(* Logix 5000 project; controller NWGG 1756-L72 rev 35.12; software revision 35.00; part 15 of 19 *)
(* tags used below, declared in another part *)
   Air_Gates_Opened : BOOL;
   ALM_Air_Gate_Failed_Open_Bin17 : ALARM_DIGITAL;
   ALM_Air_Gate_Failed_Open_Bin18 : ALARM_DIGITAL;
   ALM_Air_Gate_Failed_Open_Bin19 : ALARM_DIGITAL;
   ALM_Air_Gate_Failed_Open_Bin20 : ALARM_DIGITAL;
   ALM_Air_Gate_Failed_Open_Bin21 : ALARM_DIGITAL;
   ALM_Air_Gate_Failed_Open_Bin22 : ALARM_DIGITAL;
   ALM_Air_Gate_Failed_Open_Bin23 : ALARM_DIGITAL;
   ALM_Air_Gate_Failed_Open_Bin24 : ALARM_DIGITAL;
   ALM_Air_Gate_Failed_Open_Bin25 : ALARM_DIGITAL;
   ALM_Air_Gate_Failed_Open_Bin26 : ALARM_DIGITAL;
   ALM_Air_Gate_Failed_Open_Bin27 : ALARM_DIGITAL;
   ALM_Air_Gate_Failed_Open_Bin28 : ALARM_DIGITAL;
   Auto_Stop_Clean : BOOL;
   Belt : udt_Motor[16];
   Belts_Ready : BOOL;
   Belts_Running : BOOL;
   Bin_Clean_Pause : BOOL;
   Bin_Loadout_Control : Loadout_Bin_Control[29];
   Bin_Transfer_Pause : BOOL;
   Bin_Treat_Pause : BOOL;
   Bins_Rqd : BOOL;
   ckIDX : DINT;
   Clean_Batch_Status : DINT;
   Clean_Bin_Gates_Opened : BOOL;
   Clean_Interlock : BOOL;
   Clean_Scale_Unavailable : BOOL;
   cntCleanTime : COUNTER;
   Concrete_Clean_Belts_Ready : BOOL;
   Concrete_Leg : udt_Motor;
   Current_Dist_List_IDX : DINT;
   Current_Transfer_Bin_From : BOOL[32];
   Current_Transfer_Bin_To : BOOL[32];
   IDX : DINT;
   Loadout_Bin : udt_Loadout_Bin[29];
   Loadout_K_Valve : udt_Loadout_K_Valve[2];
   Loop_Idx : DINT;
   Manual_Mode : BOOL;
   NA : BOOL;
   Pause_Load_By_Time : BOOL[32];
   Pause_Load_By_Weight : BOOL[32];
   Pause_Load_Expired : DINT[2];
   Pause_Load_Pre : DINT[2];
   Reversing_Belt_Bypass_Valve : BOOL;
   Reversing_Belt_Reversed : BOOL;
   Start_Clean_Belts_Enabled : BOOL;
   Steel_Rqd_Belts_Running : BOOL;
   Target_Weight : DINT[2];
   TMR_Max_Clean_Delay : TIMER;
   TMR_Max_Treat_Delay : TIMER;
   tmr_Pause_Load_Timer : TIMER[2];
   tmrCleanTime : TIMER;
   Transfer_Batch_Status : DINT;
   Transfer_From_IDX : DINT;
   Transfer_To_IDX : DINT;
   Treat_Batch_Status : DINT;
   Treat_Bin_Gates_Opened : BOOL;
   Treat_Bins_Open : BOOL;
   Treat_Scale_Unavailable : BOOL;
   Use_Concrete_Side_Clean : BOOL;
   Use_Steel_Side_Clean : BOOL;
   Use_Steel_Transfer_Bins : BOOL;
   I1_000_Bit02 : ALIAS FOR I1.2;
   I1_000_Bit03 : ALIAS FOR I1.3;
   I1_000_Bit04 : ALIAS FOR I1.4;
   I1_000_Bit06 : ALIAS FOR I1.6;
   I1_000_Bit07 : ALIAS FOR I1.7;
   I1_000_Bit09 : ALIAS FOR I1.9;
   I1_000_Bit10 : ALIAS FOR I1.10;
   I1_000_Bit12 : ALIAS FOR I1.12;
   I1_000_Bit13 : ALIAS FOR I1.13;
   I1_000_Bit15 : ALIAS FOR I1.15;
   I2_000_Bit00 : ALIAS FOR I2.0;
   I2_000_Bit03 : ALIAS FOR I2.3;
   I2_000_Bit06 : ALIAS FOR I2.6;
   I2_000_Bit09 : ALIAS FOR I2.9;
   I2_000_Bit12 : ALIAS FOR I2.12;
   I3_000_Bit00 : ALIAS FOR I3.0;
   I3_000_Bit03 : ALIAS FOR I3.3;
   I3_000_Bit06 : ALIAS FOR I3.6;
   I4_000_Bit09 : ALIAS FOR I4.9;
   I4_000_Bit10 : ALIAS FOR I4.10;
   I4_000_Bit12 : ALIAS FOR I4.12;
   I4_000_Bit13 : ALIAS FOR I4.13;
   I4_000_Bit14 : ALIAS FOR I4.14;
   I4_000_Bit15 : ALIAS FOR I4.15;
   O10_000_Bit00 : ALIAS FOR O10.0;
   O10_000_Bit01 : ALIAS FOR O10.1;
   O10_000_Bit02 : ALIAS FOR O10.2;
   O10_000_Bit03 : ALIAS FOR O10.3;
   O10_000_Bit04 : ALIAS FOR O10.4;
   O10_000_Bit05 : ALIAS FOR O10.5;
   O10_000_Bit06 : ALIAS FOR O10.6;
   O10_000_Bit07 : ALIAS FOR O10.7;
   O10_000_Bit08 : ALIAS FOR O10.8;
   O10_000_Bit09 : ALIAS FOR O10.9;
   O10_000_Bit10 : ALIAS FOR O10.10;
   O10_000_Bit11 : ALIAS FOR O10.11;
   O10_000_Bit12 : ALIAS FOR O10.12;
   O10_000_Bit13 : ALIAS FOR O10.13;
   O10_000_Bit14 : ALIAS FOR O10.14;
   O11_000_Bit00 : ALIAS FOR O11.0;
   O11_000_Bit01 : ALIAS FOR O11.1;
   O11_000_Bit02 : ALIAS FOR O11.2;
   O11_000_Bit03 : ALIAS FOR O11.3;
   O11_000_Bit04 : ALIAS FOR O11.4;
   O11_000_Bit05 : ALIAS FOR O11.5;
   O11_000_Bit06 : ALIAS FOR O11.6;
   O11_000_Bit07 : ALIAS FOR O11.7;
   O11_000_Bit08 : ALIAS FOR O11.8;
   O9_000_Bit03 : ALIAS FOR O9.3;
   O9_000_Bit04 : ALIAS FOR O9.4;
   O9_000_Bit05 : ALIAS FOR O9.5;
   O9_000_Bit06 : ALIAS FOR O9.6;
   O9_000_Bit07 : ALIAS FOR O9.7;
   O9_000_Bit08 : ALIAS FOR O9.8;
   O9_000_Bit09 : ALIAS FOR O9.9;
   O9_000_Bit10 : ALIAS FOR O9.10;
   O9_000_Bit11 : ALIAS FOR O9.11;
   O9_000_Bit12 : ALIAS FOR O9.12;
   O9_000_Bit13 : ALIAS FOR O9.13;
   O9_000_Bit14 : ALIAS FOR O9.14;
   Truck_Scales : udt_Truck_Scale[2];
(* SeedLoadoutMain, continued *)

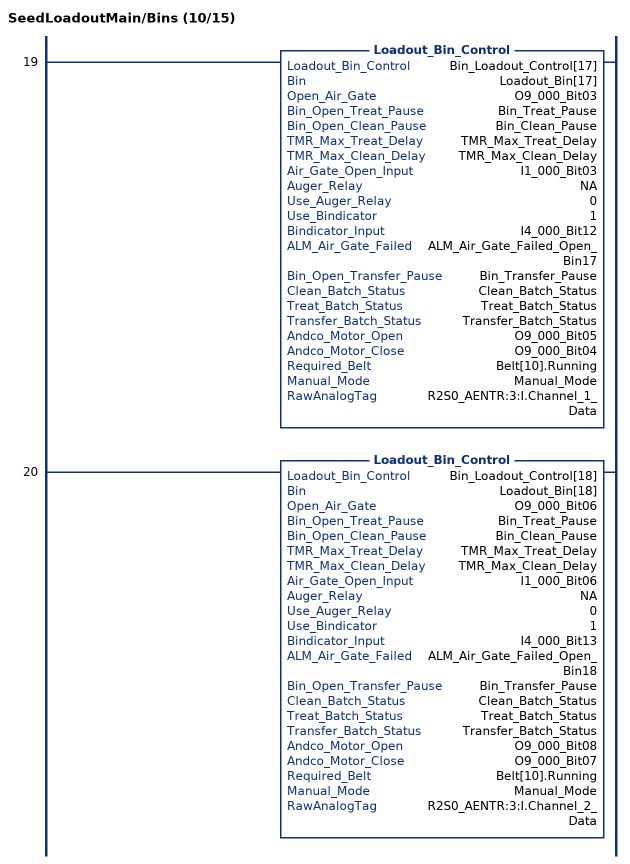
   19: Loadout_Bin_Control(Bin_Loadout_Control[17],Loadout_Bin[17],O9_000_Bit03,Bin_Treat_Pause,Bin_Clean_Pause,TMR_Max_Treat_Delay,TMR_Max_Clean_Delay,I1_000_Bit03,NA,0,1,I4_000_Bit12,ALM_Air_Gate_Failed_Open_Bin17,Bin_Transfer_Pause,Clean_Batch_Status,Treat_Batch_Status,Transfer_Batch_Status,O9_000_Bit05,O9_000_Bit04,Belt[10].Running,Manual_Mode,R2S0_AENTR:3:I.Channel_1_Data);
   20: Loadout_Bin_Control(Bin_Loadout_Control[18],Loadout_Bin[18],O9_000_Bit06,Bin_Treat_Pause,Bin_Clean_Pause,TMR_Max_Treat_Delay,TMR_Max_Clean_Delay,I1_000_Bit06,NA,0,1,I4_000_Bit13,ALM_Air_Gate_Failed_Open_Bin18,Bin_Transfer_Pause,Clean_Batch_Status,Treat_Batch_Status,Transfer_Batch_Status,O9_000_Bit08,O9_000_Bit07,Belt[10].Running,Manual_Mode,R2S0_AENTR:3:I.Channel_2_Data);
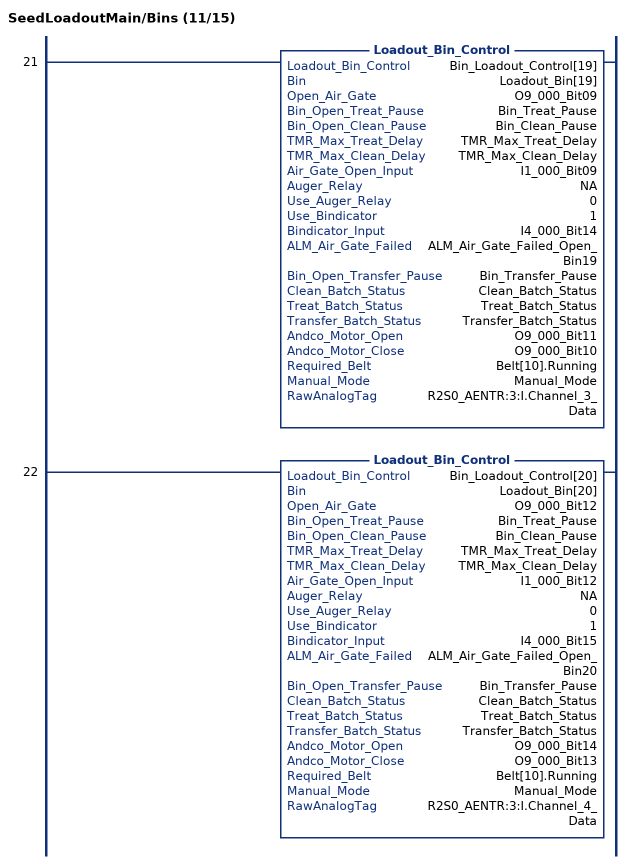
   21: Loadout_Bin_Control(Bin_Loadout_Control[19],Loadout_Bin[19],O9_000_Bit09,Bin_Treat_Pause,Bin_Clean_Pause,TMR_Max_Treat_Delay,TMR_Max_Clean_Delay,I1_000_Bit09,NA,0,1,I4_000_Bit14,ALM_Air_Gate_Failed_Open_Bin19,Bin_Transfer_Pause,Clean_Batch_Status,Treat_Batch_Status,Transfer_Batch_Status,O9_000_Bit11,O9_000_Bit10,Belt[10].Running,Manual_Mode,R2S0_AENTR:3:I.Channel_3_Data);
   22: Loadout_Bin_Control(Bin_Loadout_Control[20],Loadout_Bin[20],O9_000_Bit12,Bin_Treat_Pause,Bin_Clean_Pause,TMR_Max_Treat_Delay,TMR_Max_Clean_Delay,I1_000_Bit12,NA,0,1,I4_000_Bit15,ALM_Air_Gate_Failed_Open_Bin20,Bin_Transfer_Pause,Clean_Batch_Status,Treat_Batch_Status,Transfer_Batch_Status,O9_000_Bit14,O9_000_Bit13,Belt[10].Running,Manual_Mode,R2S0_AENTR:3:I.Channel_4_Data);
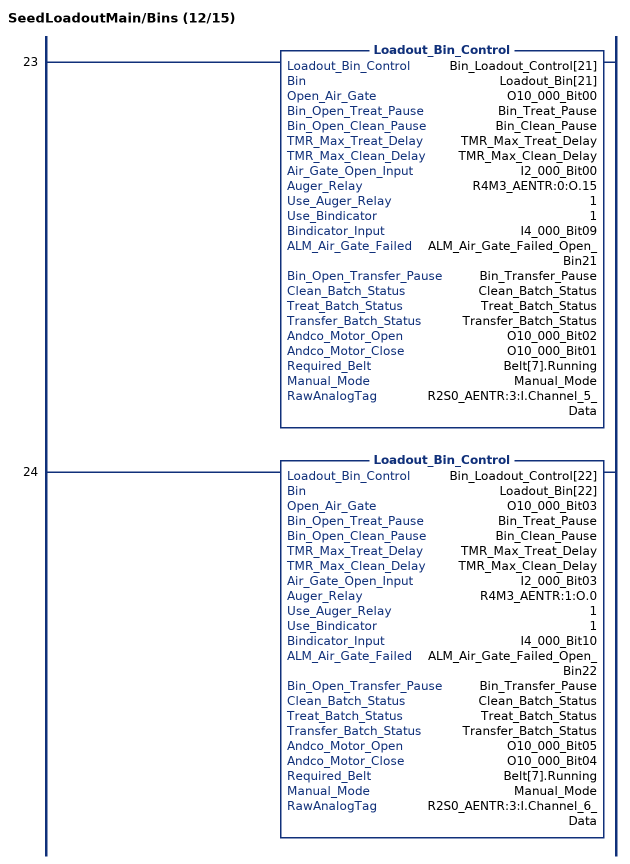
   23: Loadout_Bin_Control(Bin_Loadout_Control[21],Loadout_Bin[21],O10_000_Bit00,Bin_Treat_Pause,Bin_Clean_Pause,TMR_Max_Treat_Delay,TMR_Max_Clean_Delay,I2_000_Bit00,R4M3_AENTR:0:O.15,1,1,I4_000_Bit09,ALM_Air_Gate_Failed_Open_Bin21,Bin_Transfer_Pause,Clean_Batch_Status,Treat_Batch_Status,Transfer_Batch_Status,O10_000_Bit02,O10_000_Bit01,Belt[7].Running,Manual_Mode,R2S0_AENTR:3:I.Channel_5_Data);
   24: Loadout_Bin_Control(Bin_Loadout_Control[22],Loadout_Bin[22],O10_000_Bit03,Bin_Treat_Pause,Bin_Clean_Pause,TMR_Max_Treat_Delay,TMR_Max_Clean_Delay,I2_000_Bit03,R4M3_AENTR:1:O.0,1,1,I4_000_Bit10,ALM_Air_Gate_Failed_Open_Bin22,Bin_Transfer_Pause,Clean_Batch_Status,Treat_Batch_Status,Transfer_Batch_Status,O10_000_Bit05,O10_000_Bit04,Belt[7].Running,Manual_Mode,R2S0_AENTR:3:I.Channel_6_Data);
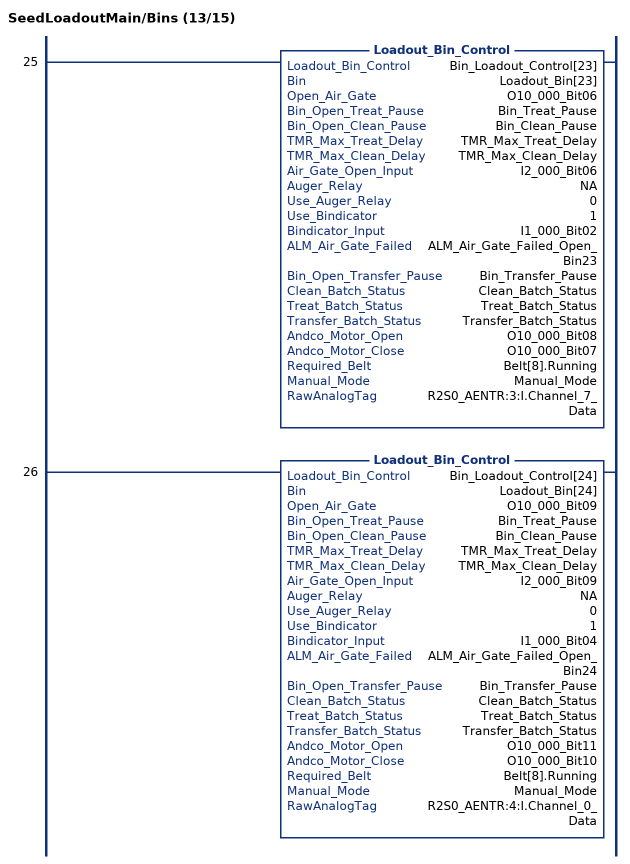
   25: Loadout_Bin_Control(Bin_Loadout_Control[23],Loadout_Bin[23],O10_000_Bit06,Bin_Treat_Pause,Bin_Clean_Pause,TMR_Max_Treat_Delay,TMR_Max_Clean_Delay,I2_000_Bit06,NA,0,1,I1_000_Bit02,ALM_Air_Gate_Failed_Open_Bin23,Bin_Transfer_Pause,Clean_Batch_Status,Treat_Batch_Status,Transfer_Batch_Status,O10_000_Bit08,O10_000_Bit07,Belt[8].Running,Manual_Mode,R2S0_AENTR:3:I.Channel_7_Data);
   26: Loadout_Bin_Control(Bin_Loadout_Control[24],Loadout_Bin[24],O10_000_Bit09,Bin_Treat_Pause,Bin_Clean_Pause,TMR_Max_Treat_Delay,TMR_Max_Clean_Delay,I2_000_Bit09,NA,0,1,I1_000_Bit04,ALM_Air_Gate_Failed_Open_Bin24,Bin_Transfer_Pause,Clean_Batch_Status,Treat_Batch_Status,Transfer_Batch_Status,O10_000_Bit11,O10_000_Bit10,Belt[8].Running,Manual_Mode,R2S0_AENTR:4:I.Channel_0_Data);
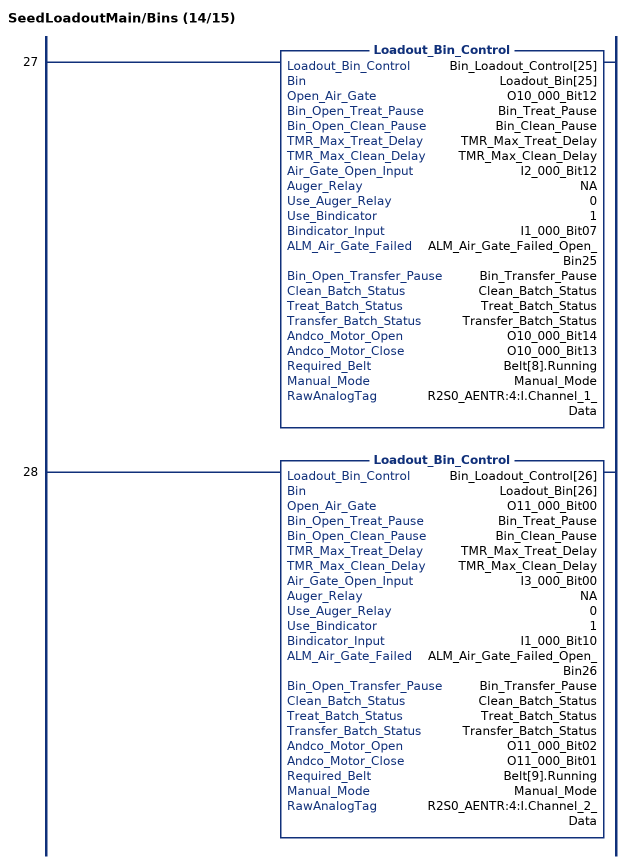
   27: Loadout_Bin_Control(Bin_Loadout_Control[25],Loadout_Bin[25],O10_000_Bit12,Bin_Treat_Pause,Bin_Clean_Pause,TMR_Max_Treat_Delay,TMR_Max_Clean_Delay,I2_000_Bit12,NA,0,1,I1_000_Bit07,ALM_Air_Gate_Failed_Open_Bin25,Bin_Transfer_Pause,Clean_Batch_Status,Treat_Batch_Status,Transfer_Batch_Status,O10_000_Bit14,O10_000_Bit13,Belt[8].Running,Manual_Mode,R2S0_AENTR:4:I.Channel_1_Data);
   28: Loadout_Bin_Control(Bin_Loadout_Control[26],Loadout_Bin[26],O11_000_Bit00,Bin_Treat_Pause,Bin_Clean_Pause,TMR_Max_Treat_Delay,TMR_Max_Clean_Delay,I3_000_Bit00,NA,0,1,I1_000_Bit10,ALM_Air_Gate_Failed_Open_Bin26,Bin_Transfer_Pause,Clean_Batch_Status,Treat_Batch_Status,Transfer_Batch_Status,O11_000_Bit02,O11_000_Bit01,Belt[9].Running,Manual_Mode,R2S0_AENTR:4:I.Channel_2_Data);
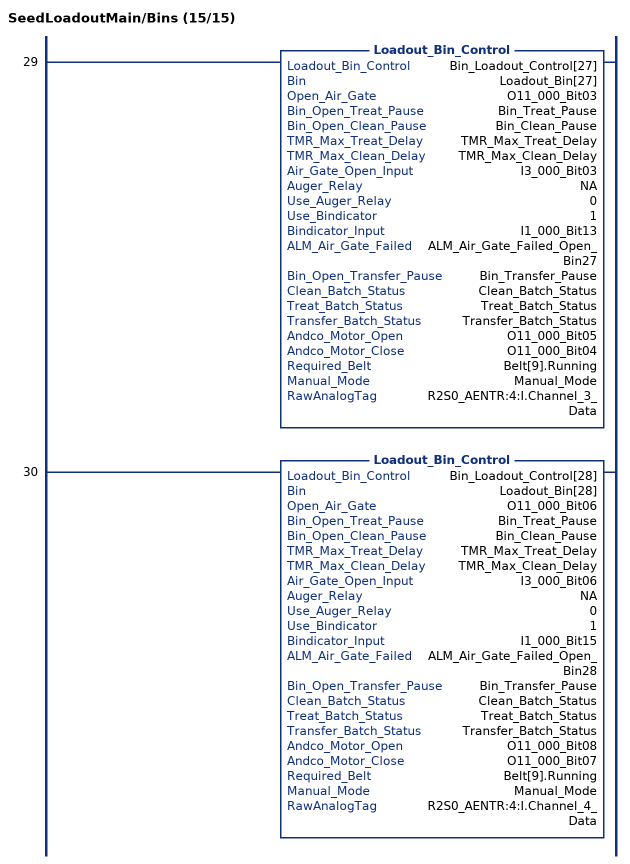
   29: Loadout_Bin_Control(Bin_Loadout_Control[27],Loadout_Bin[27],O11_000_Bit03,Bin_Treat_Pause,Bin_Clean_Pause,TMR_Max_Treat_Delay,TMR_Max_Clean_Delay,I3_000_Bit03,NA,0,1,I1_000_Bit13,ALM_Air_Gate_Failed_Open_Bin27,Bin_Transfer_Pause,Clean_Batch_Status,Treat_Batch_Status,Transfer_Batch_Status,O11_000_Bit05,O11_000_Bit04,Belt[9].Running,Manual_Mode,R2S0_AENTR:4:I.Channel_3_Data);
   30: Loadout_Bin_Control(Bin_Loadout_Control[28],Loadout_Bin[28],O11_000_Bit06,Bin_Treat_Pause,Bin_Clean_Pause,TMR_Max_Treat_Delay,TMR_Max_Clean_Delay,I3_000_Bit06,NA,0,1,I1_000_Bit15,ALM_Air_Gate_Failed_Open_Bin28,Bin_Transfer_Pause,Clean_Batch_Status,Treat_Batch_Status,Transfer_Batch_Status,O11_000_Bit08,O11_000_Bit07,Belt[9].Running,Manual_Mode,R2S0_AENTR:4:I.Channel_4_Data);
END_ROUTINE

ROUTINE Cancel_Cal_Bin   (* ladder *)
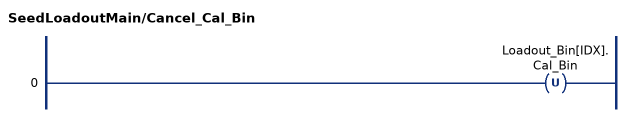
   0: OTU(Loadout_Bin[IDX].Cal_Bin);
END_ROUTINE

ROUTINE Check_Bin_Availability   (* ladder *)
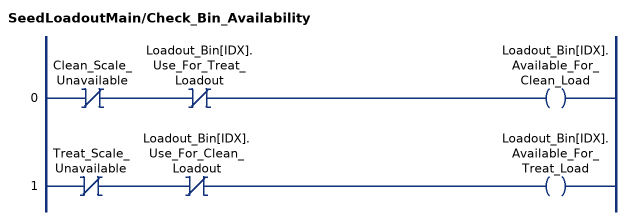
   0: XIO(Clean_Scale_Unavailable)XIO(Loadout_Bin[IDX].Use_For_Treat_Loadout)OTE(Loadout_Bin[IDX].Available_For_Clean_Load);
   1: XIO(Treat_Scale_Unavailable)XIO(Loadout_Bin[IDX].Use_For_Clean_Loadout)OTE(Loadout_Bin[IDX].Available_For_Treat_Load);
END_ROUTINE

ROUTINE Check_If_Air_Gate_Open   (* ladder *)
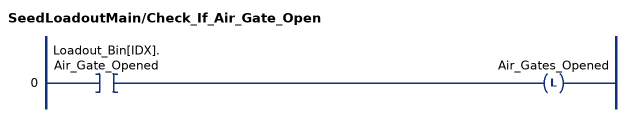
   0: XIC(Loadout_Bin[IDX].Air_Gate_Opened)OTL(Air_Gates_Opened);
END_ROUTINE

ROUTINE Check_If_Belt_Running   (* ladder *)
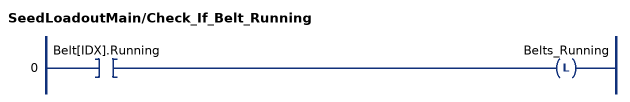
   0: XIC(Belt[IDX].Running)OTL(Belts_Running);
END_ROUTINE

ROUTINE Check_If_Treat_Gate_Open   (* ladder *)
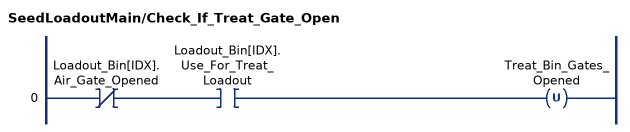
   0: XIO(Loadout_Bin[IDX].Air_Gate_Opened)XIC(Loadout_Bin[IDX].Use_For_Treat_Loadout)OTU(Treat_Bin_Gates_Opened);
END_ROUTINE

ROUTINE Check_Transfer   (* ladder *)
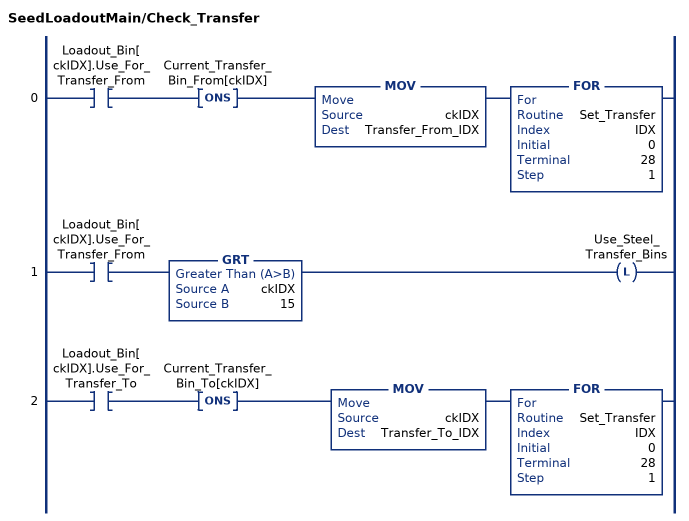
   0: XIC(Loadout_Bin[ckIDX].Use_For_Transfer_From)ONS(Current_Transfer_Bin_From[ckIDX])MOV(ckIDX,Transfer_From_IDX)FOR(Set_Transfer,IDX,0,28,1);
   1: XIC(Loadout_Bin[ckIDX].Use_For_Transfer_From)GRT(ckIDX,15)OTL(Use_Steel_Transfer_Bins);
   2: XIC(Loadout_Bin[ckIDX].Use_For_Transfer_To)ONS(Current_Transfer_Bin_To[ckIDX])MOV(ckIDX,Transfer_To_IDX)FOR(Set_Transfer,IDX,0,28,1);
END_ROUTINE

ROUTINE Check_Treater_Belts_Off   (* ladder *)
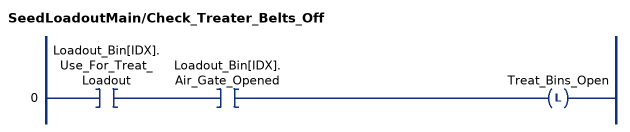
   0: XIC(Loadout_Bin[IDX].Use_For_Treat_Loadout)XIC(Loadout_Bin[IDX].Air_Gate_Opened)OTL(Treat_Bins_Open);
END_ROUTINE

ROUTINE Clean_Belt_Batch_Ready   (* ladder *)
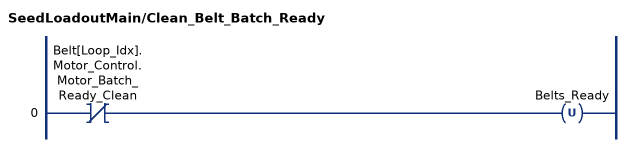
   0: XIO(Belt[Loop_Idx].Motor_Control.Motor_Batch_Ready_Clean)OTU(Belts_Ready);
END_ROUTINE

ROUTINE Clean_Belt_Start   (* ladder *)
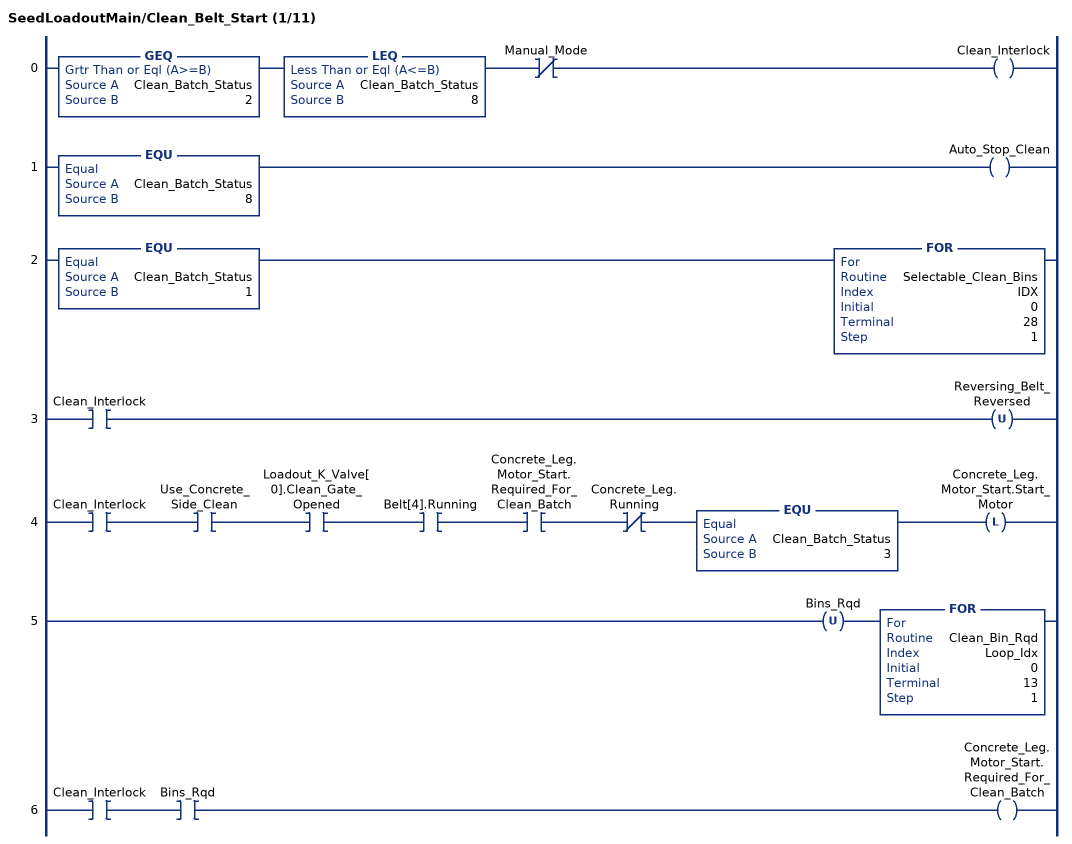
   0: GEQ(Clean_Batch_Status,2)LEQ(Clean_Batch_Status,8)XIO(Manual_Mode)OTE(Clean_Interlock);
   1: EQU(Clean_Batch_Status,8)OTE(Auto_Stop_Clean);
   2: EQU(Clean_Batch_Status,1)FOR(Selectable_Clean_Bins,IDX,0,28,1);
   3: XIC(Clean_Interlock)OTU(Reversing_Belt_Reversed);
   4: XIC(Clean_Interlock)XIC(Use_Concrete_Side_Clean)XIC(Loadout_K_Valve[0].Clean_Gate_Opened)XIC(Belt[4].Running)XIC(Concrete_Leg.Motor_Start.Required_For_Clean_Batch)XIO(Concrete_Leg.Running)EQU(Clean_Batch_Status,3)OTL(Concrete_Leg.Motor_Start.Start_Motor);
   5: OTU(Bins_Rqd)FOR(Clean_Bin_Rqd,Loop_Idx,0,13,1);
   6: XIC(Clean_Interlock)XIC(Bins_Rqd)OTE(Concrete_Leg.Motor_Start.Required_For_Clean_Batch);
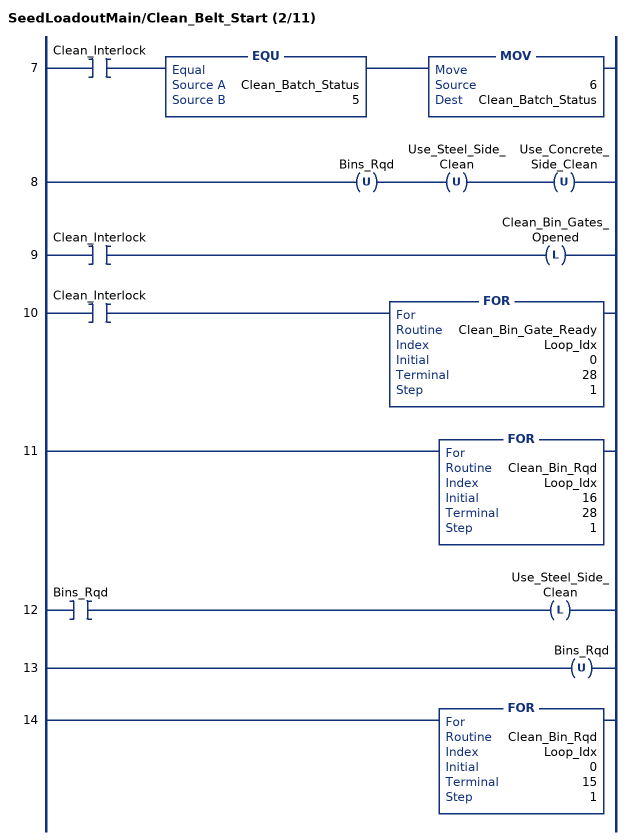
   7: XIC(Clean_Interlock)EQU(Clean_Batch_Status,5)MOV(6,Clean_Batch_Status);
   8: OTU(Bins_Rqd)OTU(Use_Steel_Side_Clean)OTU(Use_Concrete_Side_Clean);
   9: XIC(Clean_Interlock)OTL(Clean_Bin_Gates_Opened);
   10: XIC(Clean_Interlock)FOR(Clean_Bin_Gate_Ready,Loop_Idx,0,28,1);
   11: FOR(Clean_Bin_Rqd,Loop_Idx,16,28,1);
   12: XIC(Bins_Rqd)OTL(Use_Steel_Side_Clean);
   13: OTU(Bins_Rqd);
   14: FOR(Clean_Bin_Rqd,Loop_Idx,0,15,1);
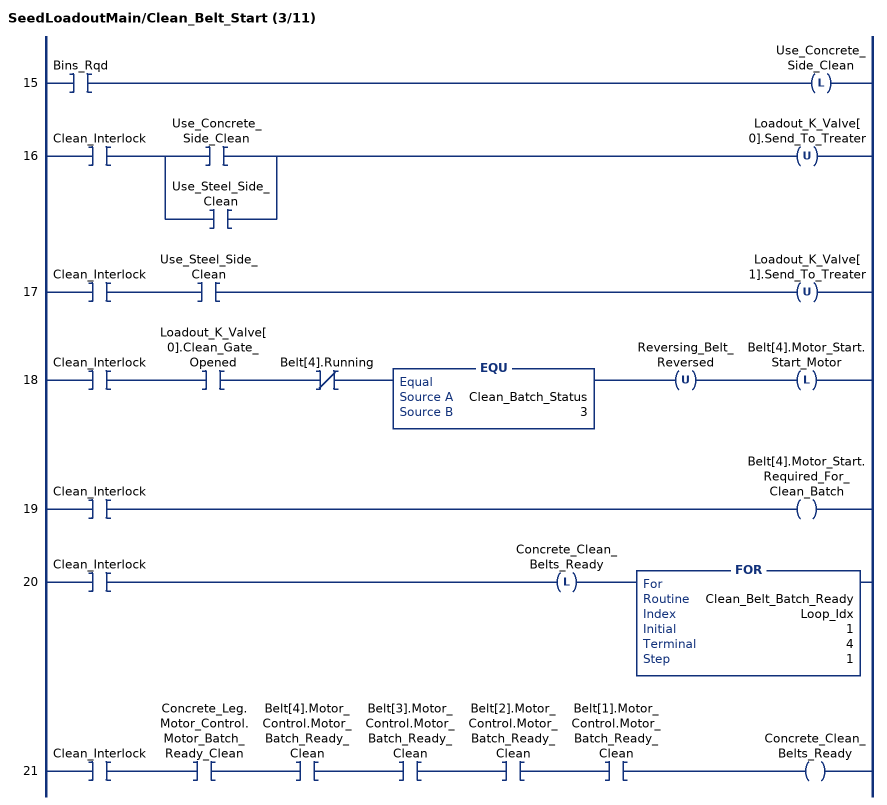
   15: XIC(Bins_Rqd)OTL(Use_Concrete_Side_Clean);
   16: XIC(Clean_Interlock)[XIC(Use_Concrete_Side_Clean) ,XIC(Use_Steel_Side_Clean) ]OTU(Loadout_K_Valve[0].Send_To_Treater);
   17: XIC(Clean_Interlock)XIC(Use_Steel_Side_Clean)OTU(Loadout_K_Valve[1].Send_To_Treater);
   18: XIC(Clean_Interlock)XIC(Loadout_K_Valve[0].Clean_Gate_Opened)XIO(Belt[4].Running)EQU(Clean_Batch_Status,3)OTU(Reversing_Belt_Reversed)OTL(Belt[4].Motor_Start.Start_Motor);
   19: XIC(Clean_Interlock)OTE(Belt[4].Motor_Start.Required_For_Clean_Batch);
   20: XIC(Clean_Interlock)OTL(Concrete_Clean_Belts_Ready)FOR(Clean_Belt_Batch_Ready,Loop_Idx,1,4,1);
   21: XIC(Clean_Interlock)XIC(Concrete_Leg.Motor_Control.Motor_Batch_Ready_Clean)XIC(Belt[4].Motor_Control.Motor_Batch_Ready_Clean)XIC(Belt[3].Motor_Control.Motor_Batch_Ready_Clean)XIC(Belt[2].Motor_Control.Motor_Batch_Ready_Clean)XIC(Belt[1].Motor_Control.Motor_Batch_Ready_Clean)OTE(Concrete_Clean_Belts_Ready);
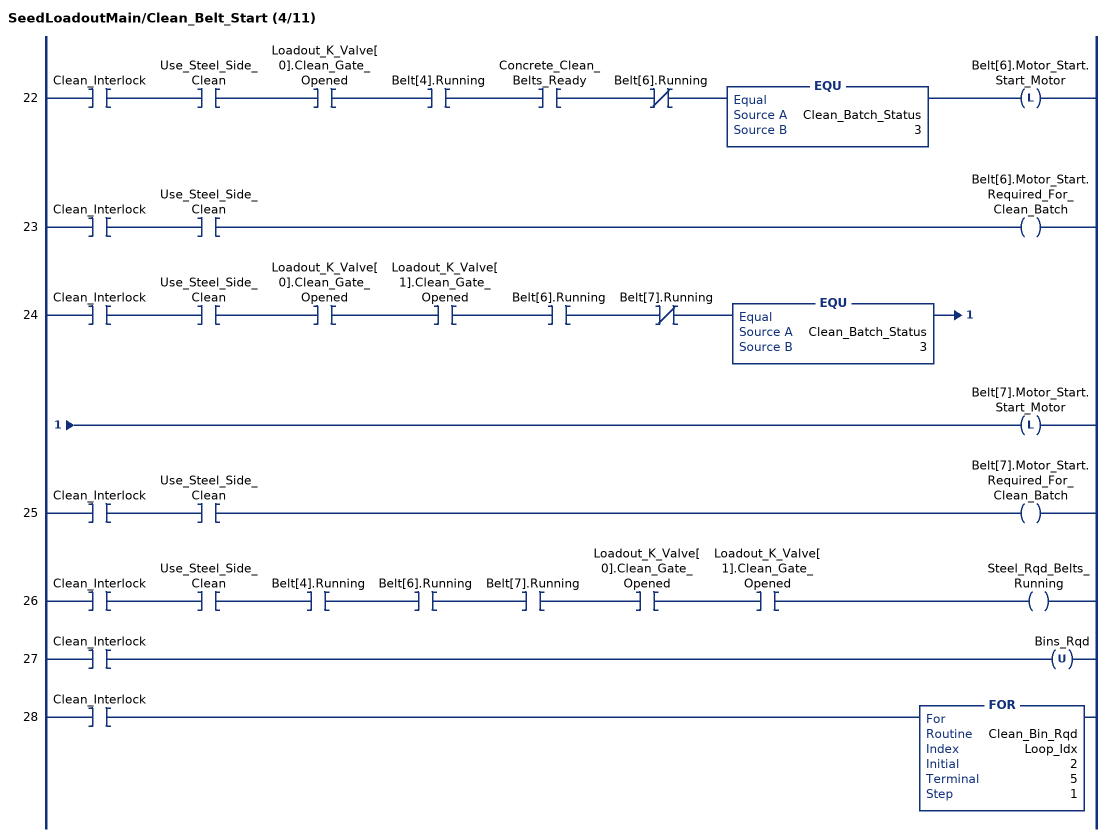
   22: XIC(Clean_Interlock)XIC(Use_Steel_Side_Clean)XIC(Loadout_K_Valve[0].Clean_Gate_Opened)XIC(Belt[4].Running)XIC(Concrete_Clean_Belts_Ready)XIO(Belt[6].Running)EQU(Clean_Batch_Status,3)OTL(Belt[6].Motor_Start.Start_Motor);
   23: XIC(Clean_Interlock)XIC(Use_Steel_Side_Clean)OTE(Belt[6].Motor_Start.Required_For_Clean_Batch);
   24: XIC(Clean_Interlock)XIC(Use_Steel_Side_Clean)XIC(Loadout_K_Valve[0].Clean_Gate_Opened)XIC(Loadout_K_Valve[1].Clean_Gate_Opened)XIC(Belt[6].Running)XIO(Belt[7].Running)EQU(Clean_Batch_Status,3)OTL(Belt[7].Motor_Start.Start_Motor);
   25: XIC(Clean_Interlock)XIC(Use_Steel_Side_Clean)OTE(Belt[7].Motor_Start.Required_For_Clean_Batch);
   26: XIC(Clean_Interlock)XIC(Use_Steel_Side_Clean)XIC(Belt[4].Running)XIC(Belt[6].Running)XIC(Belt[7].Running)XIC(Loadout_K_Valve[0].Clean_Gate_Opened)XIC(Loadout_K_Valve[1].Clean_Gate_Opened)OTE(Steel_Rqd_Belts_Running);
   27: XIC(Clean_Interlock)OTU(Bins_Rqd);
   28: XIC(Clean_Interlock)FOR(Clean_Bin_Rqd,Loop_Idx,2,5,1);
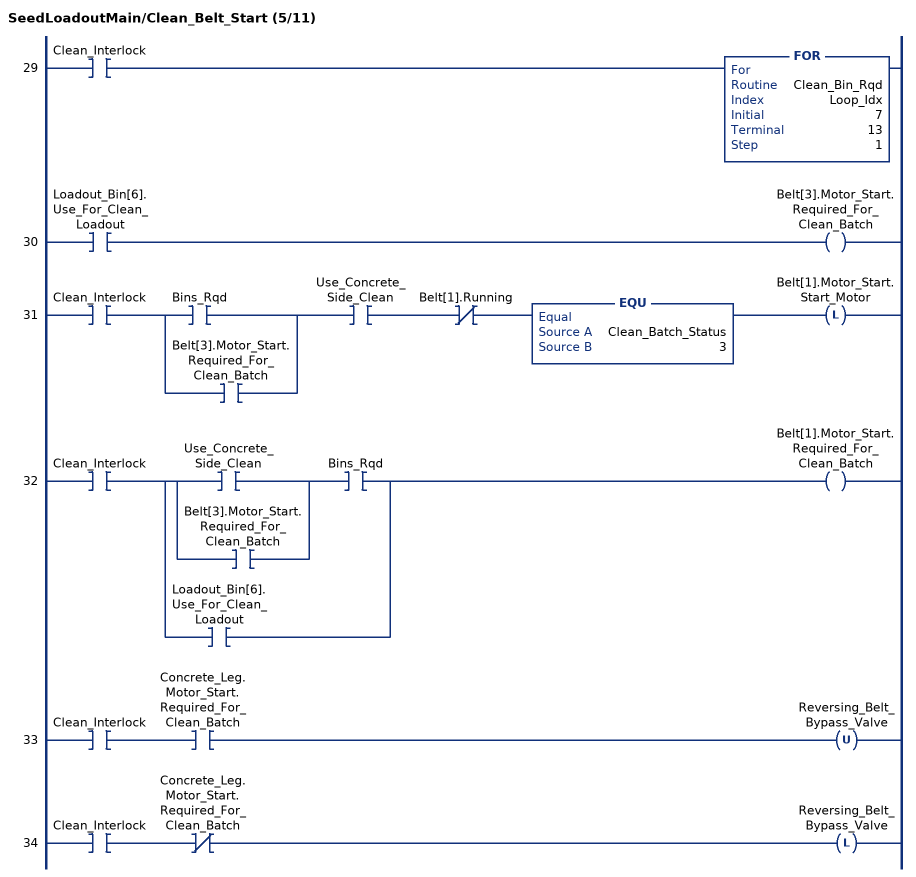
   29: XIC(Clean_Interlock)FOR(Clean_Bin_Rqd,Loop_Idx,7,13,1);
   30: XIC(Loadout_Bin[6].Use_For_Clean_Loadout)OTE(Belt[3].Motor_Start.Required_For_Clean_Batch);
   31: XIC(Clean_Interlock)[XIC(Bins_Rqd) ,XIC(Belt[3].Motor_Start.Required_For_Clean_Batch) ]XIC(Use_Concrete_Side_Clean)XIO(Belt[1].Running)EQU(Clean_Batch_Status,3)OTL(Belt[1].Motor_Start.Start_Motor);
   32: XIC(Clean_Interlock)[[XIC(Use_Concrete_Side_Clean) ,XIC(Belt[3].Motor_Start.Required_For_Clean_Batch) ] XIC(Bins_Rqd) ,XIC(Loadout_Bin[6].Use_For_Clean_Loadout) ]OTE(Belt[1].Motor_Start.Required_For_Clean_Batch);
   33: XIC(Clean_Interlock)XIC(Concrete_Leg.Motor_Start.Required_For_Clean_Batch)OTU(Reversing_Belt_Bypass_Valve);
   34: XIC(Clean_Interlock)XIO(Concrete_Leg.Motor_Start.Required_For_Clean_Batch)OTL(Reversing_Belt_Bypass_Valve);
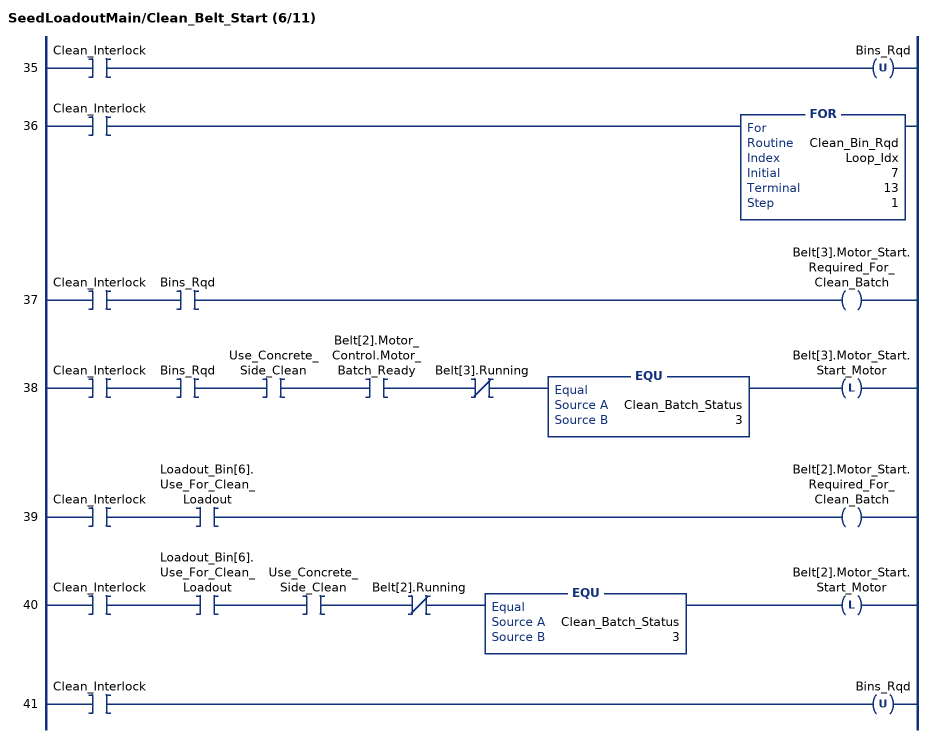
   35: XIC(Clean_Interlock)OTU(Bins_Rqd);
   36: XIC(Clean_Interlock)FOR(Clean_Bin_Rqd,Loop_Idx,7,13,1);
   37: XIC(Clean_Interlock)XIC(Bins_Rqd)OTE(Belt[3].Motor_Start.Required_For_Clean_Batch);
   38: XIC(Clean_Interlock)XIC(Bins_Rqd)XIC(Use_Concrete_Side_Clean)XIC(Belt[2].Motor_Control.Motor_Batch_Ready)XIO(Belt[3].Running)EQU(Clean_Batch_Status,3)OTL(Belt[3].Motor_Start.Start_Motor);
   39: XIC(Clean_Interlock)XIC(Loadout_Bin[6].Use_For_Clean_Loadout)OTE(Belt[2].Motor_Start.Required_For_Clean_Batch);
   40: XIC(Clean_Interlock)XIC(Loadout_Bin[6].Use_For_Clean_Loadout)XIC(Use_Concrete_Side_Clean)XIO(Belt[2].Running)EQU(Clean_Batch_Status,3)OTL(Belt[2].Motor_Start.Start_Motor);
   41: XIC(Clean_Interlock)OTU(Bins_Rqd);
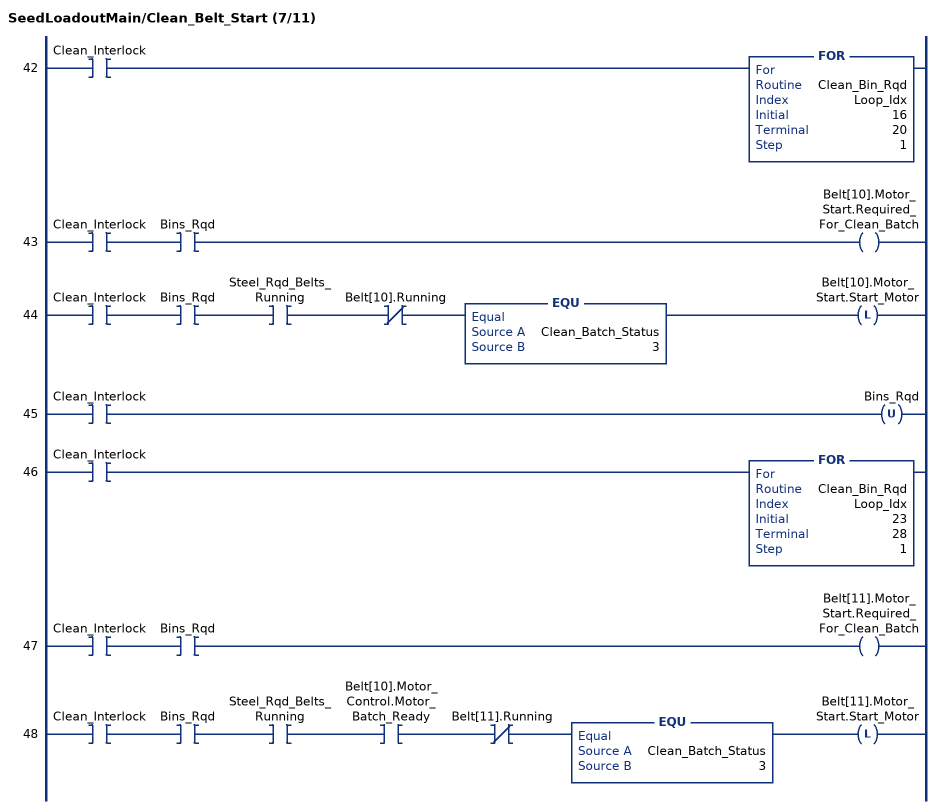
   42: XIC(Clean_Interlock)FOR(Clean_Bin_Rqd,Loop_Idx,16,20,1);
   43: XIC(Clean_Interlock)XIC(Bins_Rqd)OTE(Belt[10].Motor_Start.Required_For_Clean_Batch);
   44: XIC(Clean_Interlock)XIC(Bins_Rqd)XIC(Steel_Rqd_Belts_Running)XIO(Belt[10].Running)EQU(Clean_Batch_Status,3)OTL(Belt[10].Motor_Start.Start_Motor);
   45: XIC(Clean_Interlock)OTU(Bins_Rqd);
   46: XIC(Clean_Interlock)FOR(Clean_Bin_Rqd,Loop_Idx,23,28,1);
   47: XIC(Clean_Interlock)XIC(Bins_Rqd)OTE(Belt[11].Motor_Start.Required_For_Clean_Batch);
   48: XIC(Clean_Interlock)XIC(Bins_Rqd)XIC(Steel_Rqd_Belts_Running)XIC(Belt[10].Motor_Control.Motor_Batch_Ready)XIO(Belt[11].Running)EQU(Clean_Batch_Status,3)OTL(Belt[11].Motor_Start.Start_Motor);
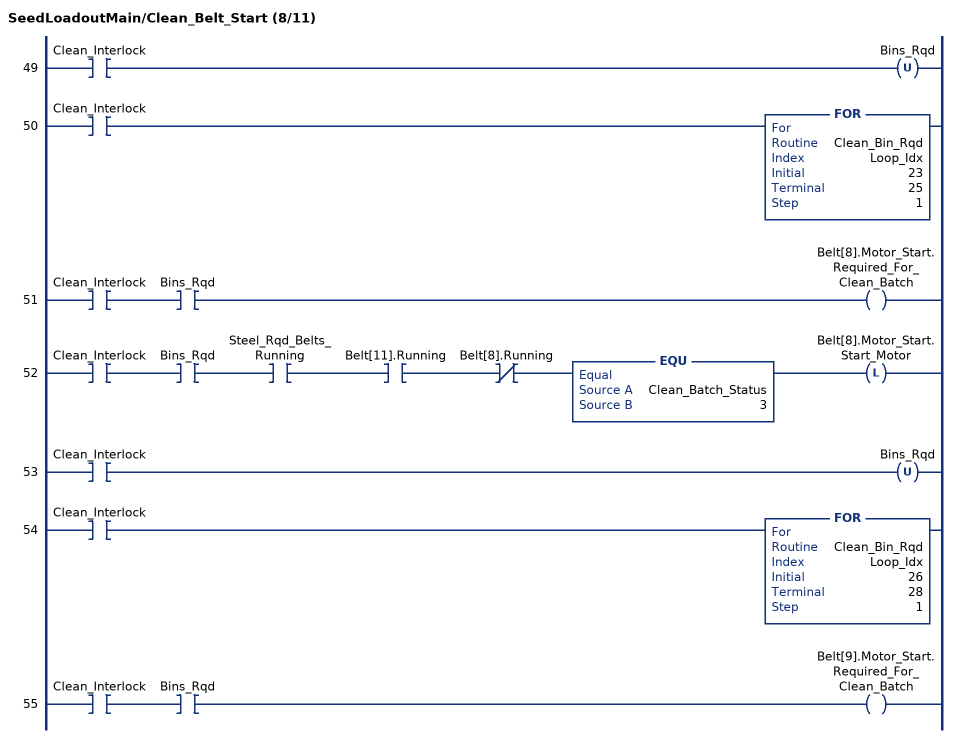
   49: XIC(Clean_Interlock)OTU(Bins_Rqd);
   50: XIC(Clean_Interlock)FOR(Clean_Bin_Rqd,Loop_Idx,23,25,1);
   51: XIC(Clean_Interlock)XIC(Bins_Rqd)OTE(Belt[8].Motor_Start.Required_For_Clean_Batch);
   52: XIC(Clean_Interlock)XIC(Bins_Rqd)XIC(Steel_Rqd_Belts_Running)XIC(Belt[11].Running)XIO(Belt[8].Running)EQU(Clean_Batch_Status,3)OTL(Belt[8].Motor_Start.Start_Motor);
   53: XIC(Clean_Interlock)OTU(Bins_Rqd);
   54: XIC(Clean_Interlock)FOR(Clean_Bin_Rqd,Loop_Idx,26,28,1);
   55: XIC(Clean_Interlock)XIC(Bins_Rqd)OTE(Belt[9].Motor_Start.Required_For_Clean_Batch);
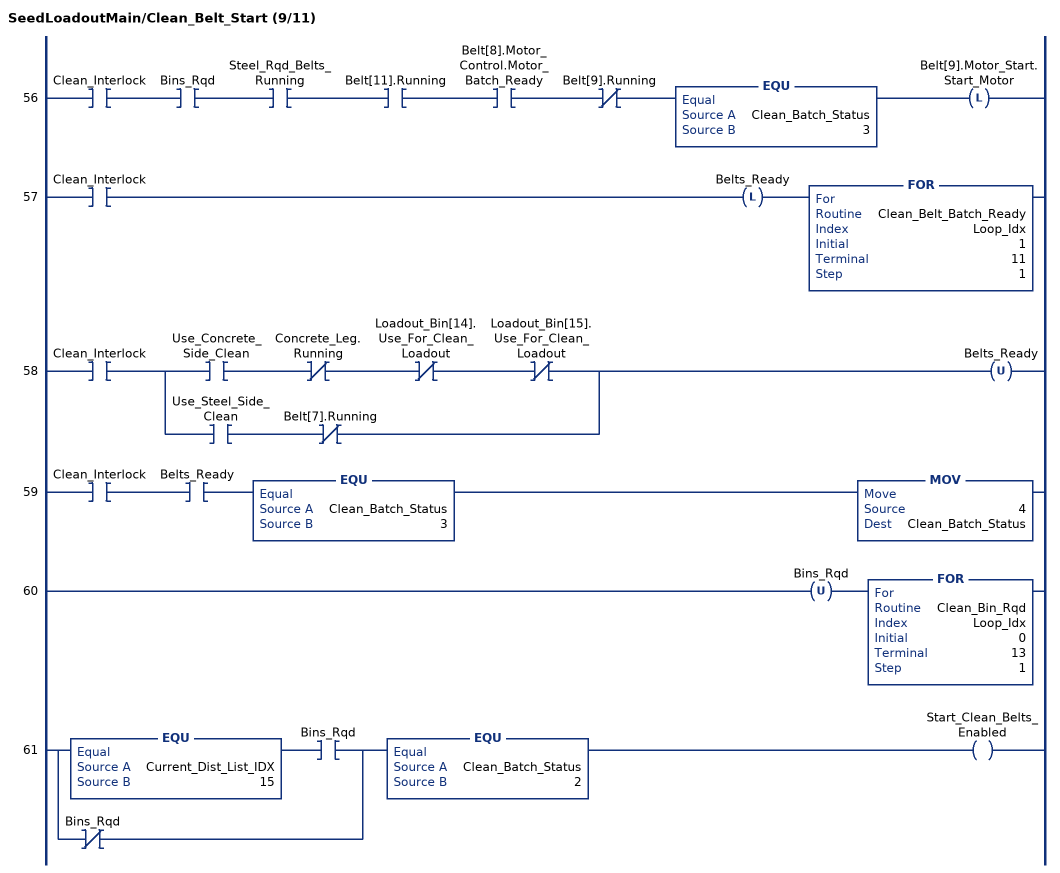
   56: XIC(Clean_Interlock)XIC(Bins_Rqd)XIC(Steel_Rqd_Belts_Running)XIC(Belt[11].Running)XIC(Belt[8].Motor_Control.Motor_Batch_Ready)XIO(Belt[9].Running)EQU(Clean_Batch_Status,3)OTL(Belt[9].Motor_Start.Start_Motor);
   57: XIC(Clean_Interlock)OTL(Belts_Ready)FOR(Clean_Belt_Batch_Ready,Loop_Idx,1,11,1);
   58: XIC(Clean_Interlock)[XIC(Use_Concrete_Side_Clean) XIO(Concrete_Leg.Running) XIO(Loadout_Bin[14].Use_For_Clean_Loadout) XIO(Loadout_Bin[15].Use_For_Clean_Loadout) ,XIC(Use_Steel_Side_Clean) XIO(Belt[7].Running) ]OTU(Belts_Ready);
   59: XIC(Clean_Interlock)XIC(Belts_Ready)EQU(Clean_Batch_Status,3)MOV(4,Clean_Batch_Status);
   60: OTU(Bins_Rqd)FOR(Clean_Bin_Rqd,Loop_Idx,0,13,1);
   61: [EQU(Current_Dist_List_IDX,15) XIC(Bins_Rqd) ,XIO(Bins_Rqd) ]EQU(Clean_Batch_Status,2)OTE(Start_Clean_Belts_Enabled);
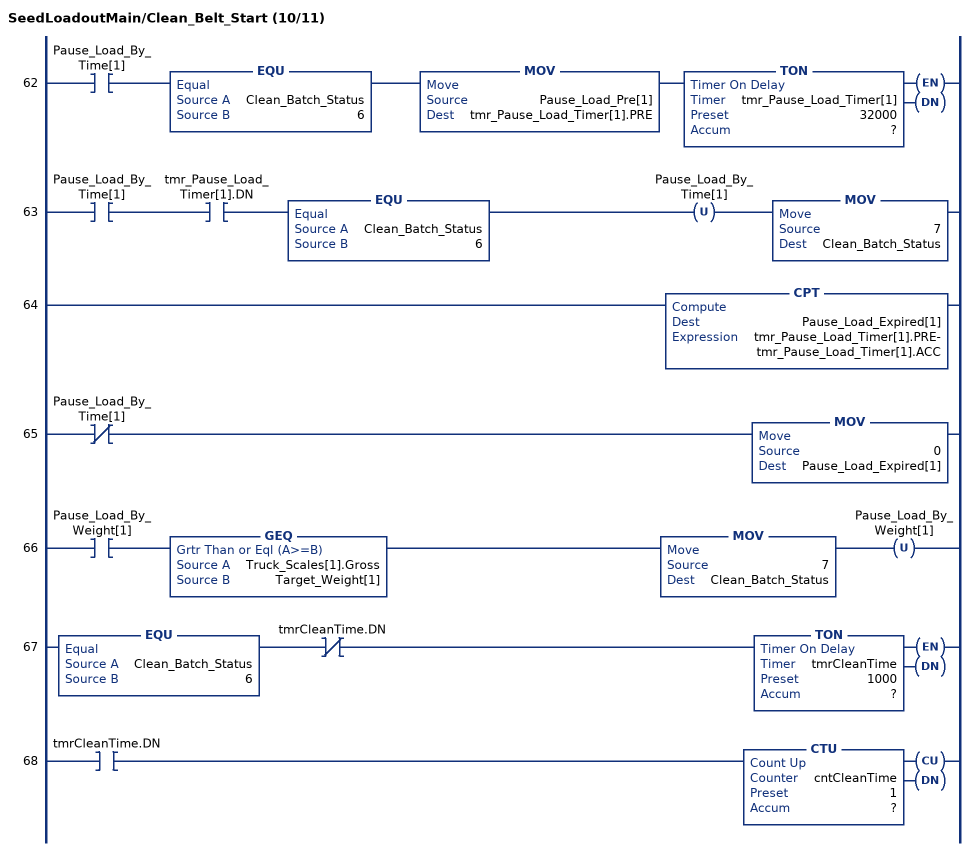
   62: XIC(Pause_Load_By_Time[1])EQU(Clean_Batch_Status,6)MOV(Pause_Load_Pre[1],tmr_Pause_Load_Timer[1].PRE)TON(tmr_Pause_Load_Timer[1],?,?);
   63: XIC(Pause_Load_By_Time[1])XIC(tmr_Pause_Load_Timer[1].DN)EQU(Clean_Batch_Status,6)OTU(Pause_Load_By_Time[1])MOV(7,Clean_Batch_Status);
   64: CPT(Pause_Load_Expired[1],tmr_Pause_Load_Timer[1].PRE-tmr_Pause_Load_Timer[1].ACC);
   65: XIO(Pause_Load_By_Time[1])MOV(0,Pause_Load_Expired[1]);
   66: XIC(Pause_Load_By_Weight[1])GEQ(Truck_Scales[1].Gross,Target_Weight[1])MOV(7,Clean_Batch_Status)OTU(Pause_Load_By_Weight[1]);
   67: EQU(Clean_Batch_Status,6)XIO(tmrCleanTime.DN)TON(tmrCleanTime,?,?);
   68: XIC(tmrCleanTime.DN)CTU(cntCleanTime,?,?);
